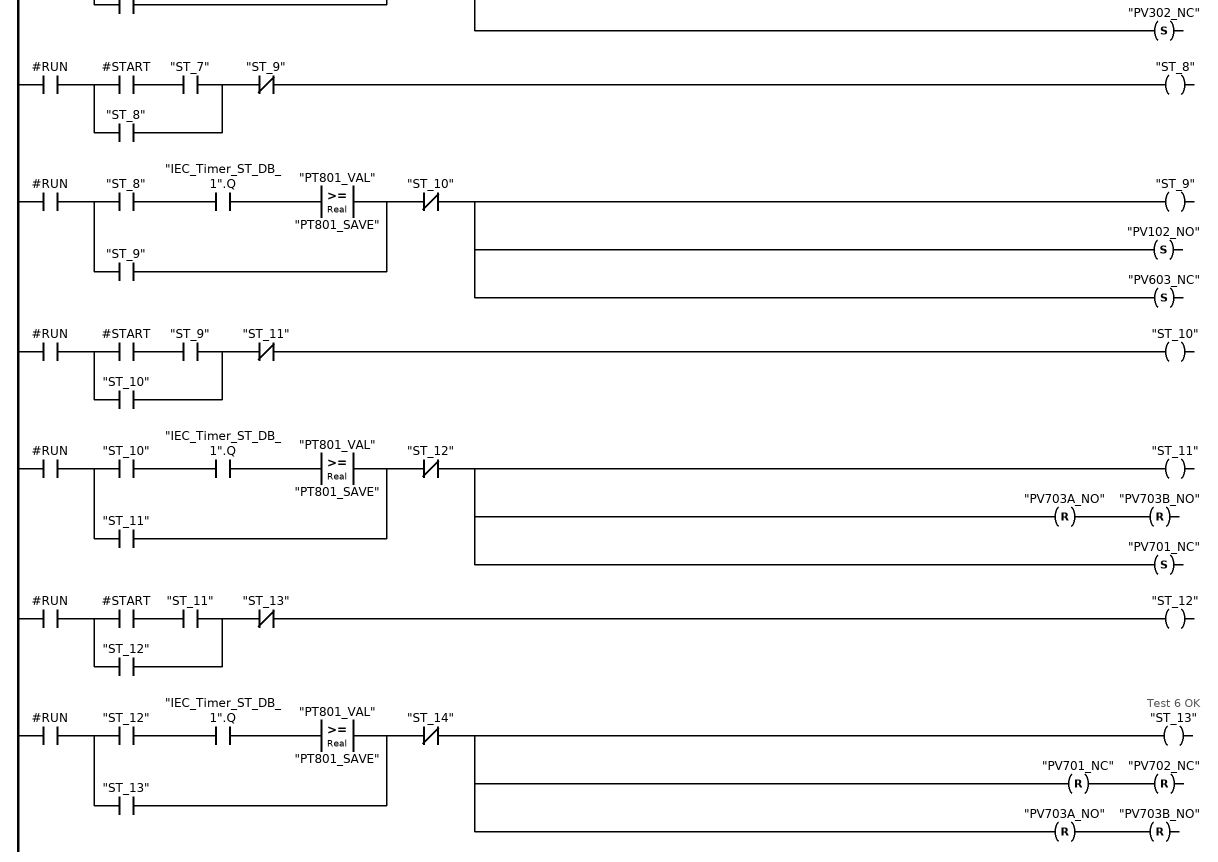
   RUNG wire#powerrail
      Contact( #RUN )
      wire#w1
      P_Contact(operand := #RUN, bit := "ST_M")
      wire#w2
      I_Contact( "ST_1" )
      I_Contact( "ST_2" )
      wire#w3
      Coil( "ST_0" )
   END_RUNG
   RUNG wire#w1
      Contact( "ST_0" )
   END_RUNG wire#w2
   RUNG wire#w3
      "ALL_VALVES_STANDBY"()
   END_RUNG
   RUNG wire#powerrail
      Contact( #RUN )
      wire#w4
      Contact( #START )
      Contact( "ST_0" )
      { S7_Templates := "SrcType := Real" } LE_Contact(in1 := "PT201_VAL", in2 := 0.0)
      { S7_Templates := "SrcType := Real" } LE_Contact(in1 := "PT401_VAL", in2 := 0.0)
      wire#w5
      I_Contact( "ST_2" )
      I_Contact( "ST_3" )
      Coil( "ST_1" )
   END_RUNG
   RUNG wire#w4
      Contact( "ST_1" )
   END_RUNG wire#w5
   RUNG wire#powerrail
      Contact( #RUN )
      wire#w6
      Contact( #START )
      Contact( "ST_1" )
      wire#w7
      I_Contact( "ST_2" )
      wire#w8
      Coil( "ST_1A" )
   END_RUNG
   RUNG wire#w6
      Contact( "ST_1A" )
   END_RUNG wire#w7
   RUNG wire#w8
      S_Coil( "PV403_NO" )
      S_Coil( "PV402_NC" )
      S_Coil( "PV602_NC" )
      S_Coil( "PV702_NC" )
   END_RUNG
   RUNG wire#w8
      Move(in := "MFC_601_MB_ADDR", out1 => "MB_DATA_MFC".MB_WRT_PARAM.MB_ADDR)
      Move(in := "MB_AD_CONTROL_MODE", out1 => "MB_DATA_MFC".MB_WRT_PARAM.DATA_ADDR)
      Move(in := "MB_VAL_CONTROL_MODE_SP_100", out1 => "MB_DATA_MFC".MB_WRT_PARAM.DATA_VAL)
   END_RUNG
   RUNG wire#powerrail
      Contact( #RUN )
      wire#w9
      Contact( "ST_1A" )
      I_Contact( "PV702_NOT_OPEN_LS" )
      wire#w10
      I_Contact( "ST_3" )
      Coil( "ST_2" )
   END_RUNG
   RUNG wire#w9
      Contact( "ST_2" )
   END_RUNG wire#w10
   RUNG wire#powerrail
      Contact( #RUN )
      wire#w11
      Contact( "ST_2" )
      Contact( "IEC_Timer_ST_DB_1".Q )
      { S7_Templates := "SrcType := Real" } GE_Contact(in1 := "PT801_VAL", in2 := "PT801_SAVE")
      wire#w12
      I_Contact( "ST_4" )
      wire#w13
      Coil( "ST_3" )
   END_RUNG
   RUNG wire#w11
      Contact( "ST_3" )
   END_RUNG wire#w12
   RUNG wire#w13
      S_Coil( "PV503_NO" )
   END_RUNG
   RUNG wire#w13
      S_Coil( "PV502_NC" )
   END_RUNG
   RUNG wire#powerrail
      Contact( #RUN )
      wire#w14
      Contact( #START )
      Contact( "ST_3" )
      wire#w15
      I_Contact( "ST_5" )
      Coil( "ST_4" )
   END_RUNG
   RUNG wire#w14
      Contact( "ST_4" )
   END_RUNG wire#w15
   RUNG wire#powerrail
      Contact( #RUN )
      wire#w16
      Contact( "ST_4" )
      Contact( "IEC_Timer_ST_DB_1".Q )
      { S7_Templates := "SrcType := Real" } GE_Contact(in1 := "PT801_VAL", in2 := "PT801_SAVE")
      wire#w17
      I_Contact( "ST_6" )
      wire#w18
      Coil( "ST_5" )
   END_RUNG
   RUNG wire#w16
      Contact( "ST_5" )
   END_RUNG wire#w17
   RUNG wire#w18
      S_Coil( "PV203_NO" )
   END_RUNG
   RUNG wire#w18
      S_Coil( "PV202_NC" )
      S_Coil( "PV601_NC" )
   END_RUNG
   RUNG wire#powerrail
      Contact( #RUN )
      wire#w19
      Contact( #START )
      Contact( "ST_5" )
      wire#w20
      I_Contact( "ST_7" )
      Coil( "ST_6" )
   END_RUNG
   RUNG wire#w19
      Contact( "ST_6" )
   END_RUNG wire#w20
   RUNG wire#powerrail
      Contact( #RUN )
      wire#w21
      Contact( "ST_6" )
      Contact( "IEC_Timer_ST_DB_1".Q )
      { S7_Templates := "SrcType := Real" } GE_Contact(in1 := "PT801_VAL", in2 := "PT801_SAVE")
      wire#w22
      I_Contact( "ST_8" )
      wire#w23
      Coil( "ST_7" )
   END_RUNG
   RUNG wire#w21
      Contact( "ST_7" )
   END_RUNG wire#w22
   RUNG wire#w23
      S_Coil( "PV303_NO" )
   END_RUNG
   RUNG wire#w23
      S_Coil( "PV302_NC" )
   END_RUNG
   RUNG wire#powerrail
      Contact( #RUN )
      wire#w24
      Contact( #START )
      Contact( "ST_7" )
      wire#w25
      I_Contact( "ST_9" )
      Coil( "ST_8" )
   END_RUNG
   RUNG wire#w24
      Contact( "ST_8" )
   END_RUNG wire#w25
   RUNG wire#powerrail
      Contact( #RUN )
      wire#w26
      Contact( "ST_8" )
      Contact( "IEC_Timer_ST_DB_1".Q )
      { S7_Templates := "SrcType := Real" } GE_Contact(in1 := "PT801_VAL", in2 := "PT801_SAVE")
      wire#w27
      I_Contact( "ST_10" )
      wire#w28
      Coil( "ST_9" )
   END_RUNG
   RUNG wire#w26
      Contact( "ST_9" )
   END_RUNG wire#w27
   RUNG wire#w28
      S_Coil( "PV102_NO" )
   END_RUNG
   RUNG wire#w28
      S_Coil( "PV603_NC" )
   END_RUNG
   RUNG wire#powerrail
      Contact( #RUN )
      wire#w29
      Contact( #START )
      Contact( "ST_9" )
      wire#w30
      I_Contact( "ST_11" )
      Coil( "ST_10" )
   END_RUNG
   RUNG wire#w29
      Contact( "ST_10" )
   END_RUNG wire#w30
   RUNG wire#powerrail
      Contact( #RUN )
      wire#w31
      Contact( "ST_10" )
      Contact( "IEC_Timer_ST_DB_1".Q )
      { S7_Templates := "SrcType := Real" } GE_Contact(in1 := "PT801_VAL", in2 := "PT801_SAVE")
      wire#w32
      I_Contact( "ST_12" )
      wire#w33
      Coil( "ST_11" )
   END_RUNG
   RUNG wire#w31
      Contact( "ST_11" )
   END_RUNG wire#w32
   RUNG wire#w33
      R_Coil( "PV703A_NO" )
      R_Coil( "PV703B_NO" )
   END_RUNG
   RUNG wire#w33
      S_Coil( "PV701_NC" )
   END_RUNG
   RUNG wire#powerrail
      Contact( #RUN )
      wire#w34
      Contact( #START )
      Contact( "ST_11" )
      wire#w35
      I_Contact( "ST_13" )
      Coil( "ST_12" )
   END_RUNG
   RUNG wire#w34
      Contact( "ST_12" )
   END_RUNG wire#w35
   RUNG wire#powerrail
      Contact( #RUN )
      wire#w36
      Contact( "ST_12" )
      Contact( "IEC_Timer_ST_DB_1".Q )
      { S7_Templates := "SrcType := Real" } GE_Contact(in1 := "PT801_VAL", in2 := "PT801_SAVE")
      wire#w37
      I_Contact( "ST_14" )
      wire#w38
      Coil( "ST_13" )   // Test 6 OK
   END_RUNG
   RUNG wire#w36
      Contact( "ST_13" )
   END_RUNG wire#w37
   RUNG wire#w38
      R_Coil( "PV701_NC" )
      R_Coil( "PV702_NC" )
   END_RUNG
   RUNG wire#w38
      R_Coil( "PV703A_NO" )
      R_Coil( "PV703B_NO" )
   END_RUNG
   // the same network as SCL:
   #_w1 := #RUN AND #RUN AND NOT "ST_M";   // rising edge of #RUN
   "ST_M" := #RUN;
   "ST_0" := (#_w1 OR (#RUN AND "ST_0")) AND NOT "ST_1" AND NOT "ST_2";
   IF "ST_0" THEN "ALL_VALVES_STANDBY"(); END_IF;
   "ST_1" := #RUN AND ((#START AND "ST_0" AND ("PT201_VAL" <= 0.0) AND ("PT401_VAL" <= 0.0)) OR "ST_1") AND NOT "ST_2" AND NOT "ST_3";
   "ST_1A" := #RUN AND ((#START AND "ST_1") OR "ST_1A") AND NOT "ST_2";
   IF "ST_1A" THEN
       "PV403_NO" := TRUE;
       "PV402_NC" := TRUE;
       "PV602_NC" := TRUE;
       "PV702_NC" := TRUE;
       "MB_DATA_MFC".MB_WRT_PARAM.MB_ADDR := "MFC_601_MB_ADDR";
       "MB_DATA_MFC".MB_WRT_PARAM.DATA_ADDR := "MB_AD_CONTROL_MODE";
       "MB_DATA_MFC".MB_WRT_PARAM.DATA_VAL := "MB_VAL_CONTROL_MODE_SP_100";
   END_IF;
   "ST_2" := #RUN AND (("ST_1A" AND NOT "PV702_NOT_OPEN_LS") OR "ST_2") AND NOT "ST_3";
   "ST_3" := #RUN AND (("ST_2" AND "IEC_Timer_ST_DB_1".Q AND ("PT801_VAL" >= "PT801_SAVE")) OR "ST_3") AND NOT "ST_4";
   IF "ST_3" THEN
       "PV503_NO" := TRUE;
       "PV502_NC" := TRUE;
   END_IF;
   "ST_4" := #RUN AND ((#START AND "ST_3") OR "ST_4") AND NOT "ST_5";
   "ST_5" := #RUN AND (("ST_4" AND "IEC_Timer_ST_DB_1".Q AND ("PT801_VAL" >= "PT801_SAVE")) OR "ST_5") AND NOT "ST_6";
   IF "ST_5" THEN
       "PV203_NO" := TRUE;
       "PV202_NC" := TRUE;
       "PV601_NC" := TRUE;
   END_IF;
   "ST_6" := #RUN AND ((#START AND "ST_5") OR "ST_6") AND NOT "ST_7";
   "ST_7" := #RUN AND (("ST_6" AND "IEC_Timer_ST_DB_1".Q AND ("PT801_VAL" >= "PT801_SAVE")) OR "ST_7") AND NOT "ST_8";
   IF "ST_7" THEN
       "PV303_NO" := TRUE;
       "PV302_NC" := TRUE;
   END_IF;
   "ST_8" := #RUN AND ((#START AND "ST_7") OR "ST_8") AND NOT "ST_9";
   "ST_9" := #RUN AND (("ST_8" AND "IEC_Timer_ST_DB_1".Q AND ("PT801_VAL" >= "PT801_SAVE")) OR "ST_9") AND NOT "ST_10";
   IF "ST_9" THEN
       "PV102_NO" := TRUE;
       "PV603_NC" := TRUE;
   END_IF;
   "ST_10" := #RUN AND ((#START AND "ST_9") OR "ST_10") AND NOT "ST_11";
   "ST_11" := #RUN AND (("ST_10" AND "IEC_Timer_ST_DB_1".Q AND ("PT801_VAL" >= "PT801_SAVE")) OR "ST_11") AND NOT "ST_12";
   IF "ST_11" THEN
       "PV703A_NO" := FALSE;
       "PV703B_NO" := FALSE;
       "PV701_NC" := TRUE;
   END_IF;
   "ST_12" := #RUN AND ((#START AND "ST_11") OR "ST_12") AND NOT "ST_13";
   "ST_13" := #RUN AND (("ST_12" AND "IEC_Timer_ST_DB_1".Q AND ("PT801_VAL" >= "PT801_SAVE")) OR "ST_13") AND NOT "ST_14";   // Test 6 OK
   IF "ST_13" THEN
       "PV701_NC" := FALSE;
       "PV702_NC" := FALSE;
       "PV703A_NO" := FALSE;
       "PV703B_NO" := FALSE;
   END_IF;
END_REGION

REGION Network 3: Process Tests
   // Tests Process Circuits  (Test #7-#9)
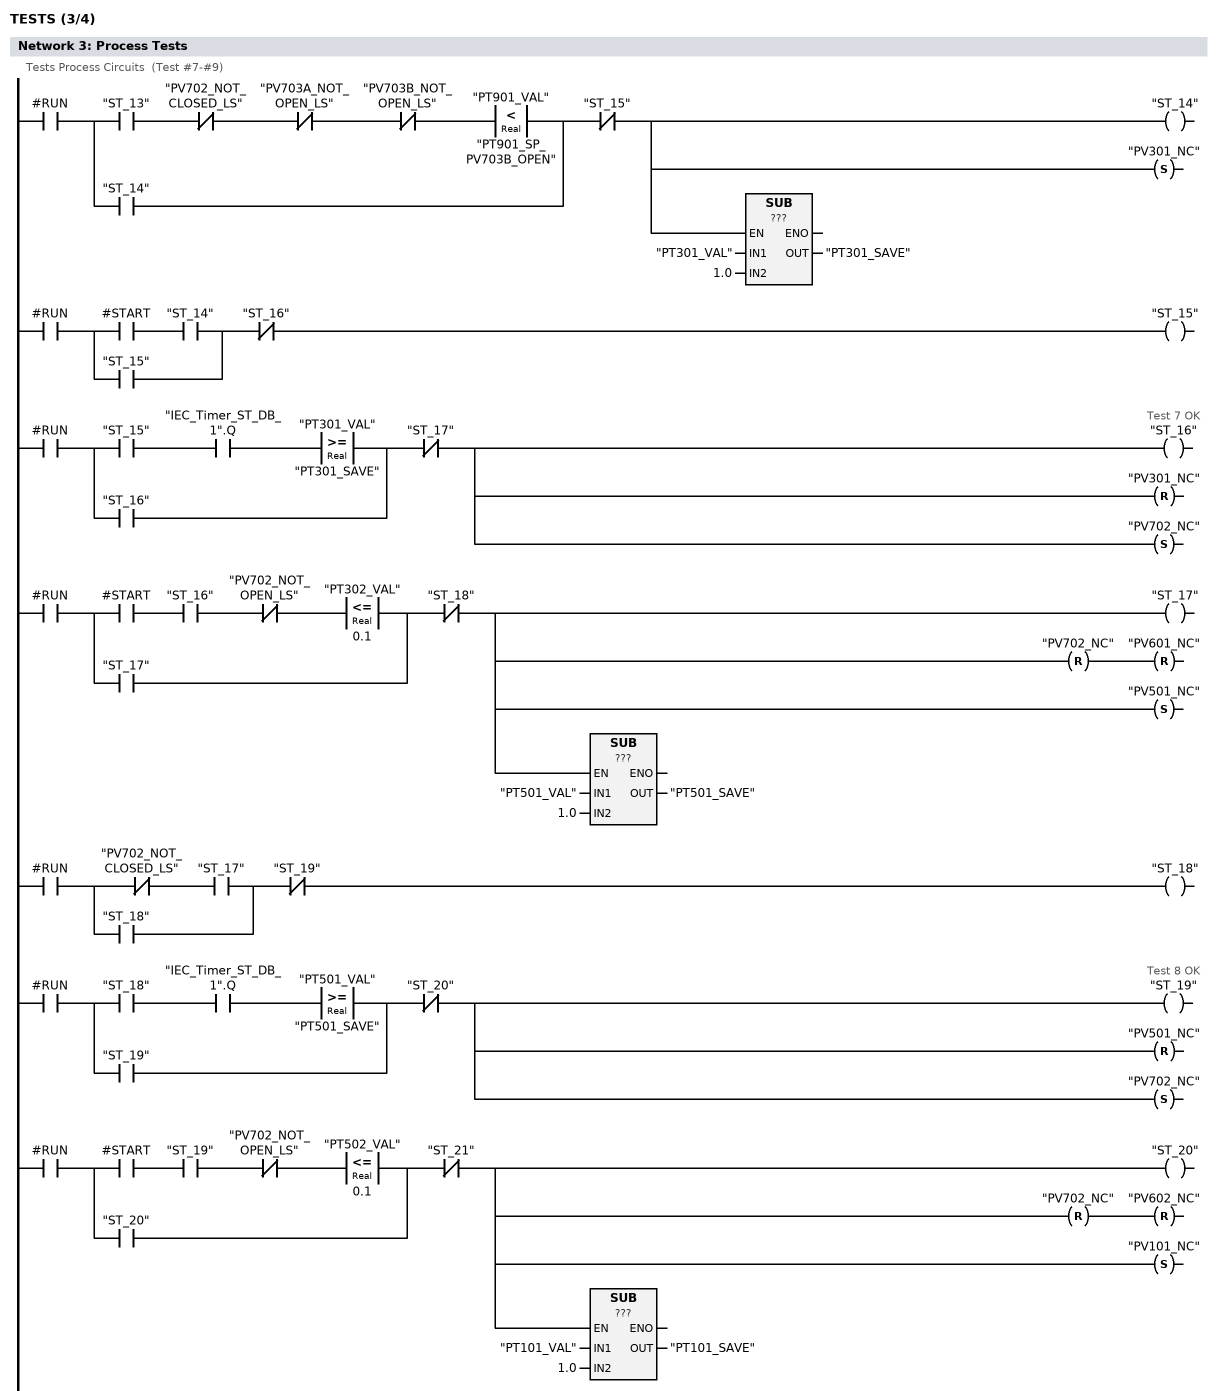
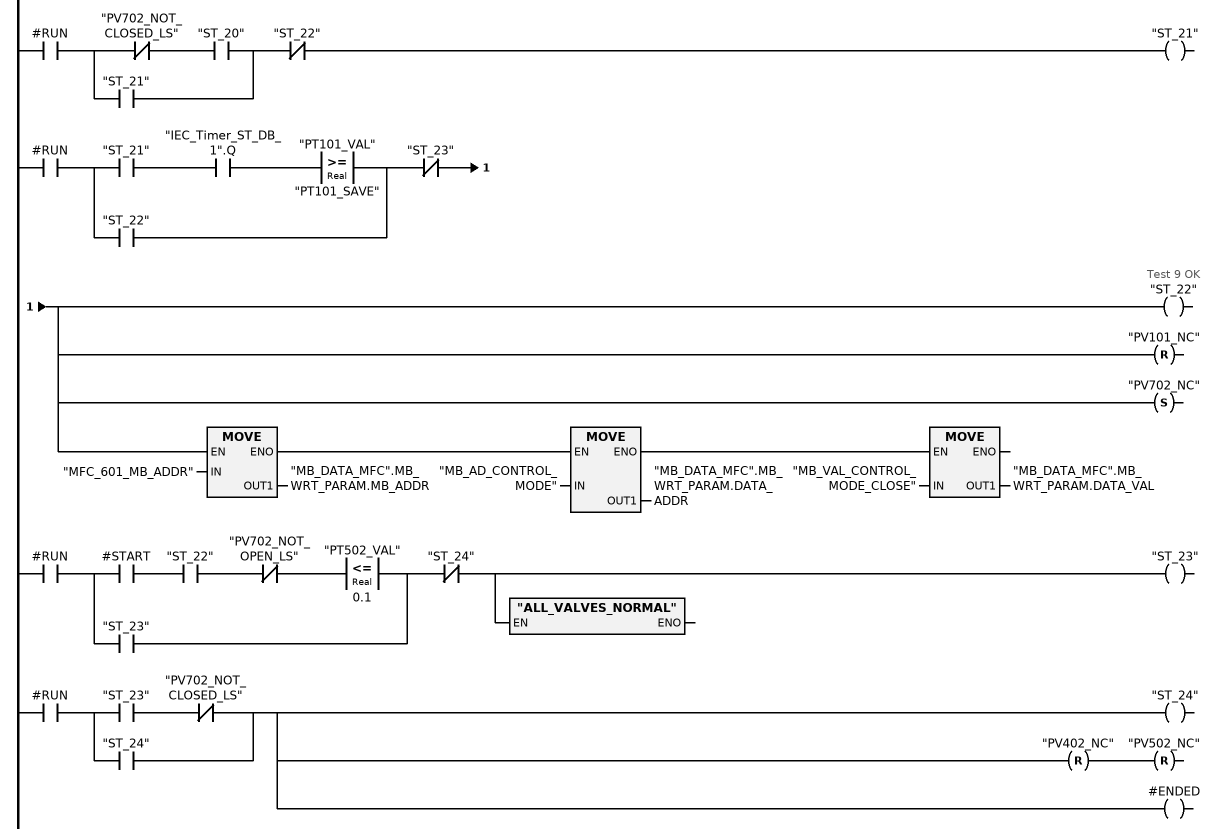
   RUNG wire#powerrail
      Contact( #RUN )
      wire#w1
      Contact( "ST_13" )
      I_Contact( "PV702_NOT_CLOSED_LS" )
      I_Contact( "PV703A_NOT_OPEN_LS" )
      I_Contact( "PV703B_NOT_OPEN_LS" )
      { S7_Templates := "SrcType := Real" } LT_Contact(in1 := "PT901_VAL", in2 := "PT901_SP_PV703B_OPEN")
      wire#w2
      I_Contact( "ST_15" )
      wire#w3
      Coil( "ST_14" )
   END_RUNG
   RUNG wire#w1
      Contact( "ST_14" )
   END_RUNG wire#w2
   RUNG wire#w3
      S_Coil( "PV301_NC" )
   END_RUNG
   RUNG wire#w3
      { S7_Templates := "SrcType := ???" } Sub(in1 := "PT301_VAL", in2 := 1.0, out => "PT301_SAVE")
   END_RUNG
   RUNG wire#powerrail
      Contact( #RUN )
      wire#w4
      Contact( #START )
      Contact( "ST_14" )
      wire#w5
      I_Contact( "ST_16" )
      Coil( "ST_15" )
   END_RUNG
   RUNG wire#w4
      Contact( "ST_15" )
   END_RUNG wire#w5
   RUNG wire#powerrail
      Contact( #RUN )
      wire#w6
      Contact( "ST_15" )
      Contact( "IEC_Timer_ST_DB_1".Q )
      { S7_Templates := "SrcType := Real" } GE_Contact(in1 := "PT301_VAL", in2 := "PT301_SAVE")
      wire#w7
      I_Contact( "ST_17" )
      wire#w8
      Coil( "ST_16" )   // Test 7 OK
   END_RUNG
   RUNG wire#w6
      Contact( "ST_16" )
   END_RUNG wire#w7
   RUNG wire#w8
      R_Coil( "PV301_NC" )
   END_RUNG
   RUNG wire#w8
      S_Coil( "PV702_NC" )
   END_RUNG
   RUNG wire#powerrail
      Contact( #RUN )
      wire#w9
      Contact( #START )
      Contact( "ST_16" )
      I_Contact( "PV702_NOT_OPEN_LS" )
      { S7_Templates := "SrcType := Real" } LE_Contact(in1 := "PT302_VAL", in2 := 0.1)
      wire#w10
      I_Contact( "ST_18" )
      wire#w11
      Coil( "ST_17" )
   END_RUNG
   RUNG wire#w9
      Contact( "ST_17" )
   END_RUNG wire#w10
   RUNG wire#w11
      R_Coil( "PV702_NC" )
      R_Coil( "PV601_NC" )
   END_RUNG
   RUNG wire#w11
      S_Coil( "PV501_NC" )
   END_RUNG
   RUNG wire#w11
      { S7_Templates := "SrcType := ???" } Sub(in1 := "PT501_VAL", in2 := 1.0, out => "PT501_SAVE")
   END_RUNG
   RUNG wire#powerrail
      Contact( #RUN )
      wire#w12
      I_Contact( "PV702_NOT_CLOSED_LS" )
      Contact( "ST_17" )
      wire#w13
      I_Contact( "ST_19" )
      Coil( "ST_18" )
   END_RUNG
   RUNG wire#w12
      Contact( "ST_18" )
   END_RUNG wire#w13
   RUNG wire#powerrail
      Contact( #RUN )
      wire#w14
      Contact( "ST_18" )
      Contact( "IEC_Timer_ST_DB_1".Q )
      { S7_Templates := "SrcType := Real" } GE_Contact(in1 := "PT501_VAL", in2 := "PT501_SAVE")
      wire#w15
      I_Contact( "ST_20" )
      wire#w16
      Coil( "ST_19" )   // Test 8 OK
   END_RUNG
   RUNG wire#w14
      Contact( "ST_19" )
   END_RUNG wire#w15
   RUNG wire#w16
      R_Coil( "PV501_NC" )
   END_RUNG
   RUNG wire#w16
      S_Coil( "PV702_NC" )
   END_RUNG
   RUNG wire#powerrail
      Contact( #RUN )
      wire#w17
      Contact( #START )
      Contact( "ST_19" )
      I_Contact( "PV702_NOT_OPEN_LS" )
      { S7_Templates := "SrcType := Real" } LE_Contact(in1 := "PT502_VAL", in2 := 0.1)
      wire#w18
      I_Contact( "ST_21" )
      wire#w19
      Coil( "ST_20" )
   END_RUNG
   RUNG wire#w17
      Contact( "ST_20" )
   END_RUNG wire#w18
   RUNG wire#w19
      R_Coil( "PV702_NC" )
      R_Coil( "PV602_NC" )
   END_RUNG
   RUNG wire#w19
      S_Coil( "PV101_NC" )
   END_RUNG
   RUNG wire#w19
      { S7_Templates := "SrcType := ???" } Sub(in1 := "PT101_VAL", in2 := 1.0, out => "PT101_SAVE")
   END_RUNG
   RUNG wire#powerrail
      Contact( #RUN )
      wire#w20
      I_Contact( "PV702_NOT_CLOSED_LS" )
      Contact( "ST_20" )
      wire#w21
      I_Contact( "ST_22" )
      Coil( "ST_21" )
   END_RUNG
   RUNG wire#w20
      Contact( "ST_21" )
   END_RUNG wire#w21
   RUNG wire#powerrail
      Contact( #RUN )
      wire#w22
      Contact( "ST_21" )
      Contact( "IEC_Timer_ST_DB_1".Q )
      { S7_Templates := "SrcType := Real" } GE_Contact(in1 := "PT101_VAL", in2 := "PT101_SAVE")
      wire#w23
      I_Contact( "ST_23" )
      wire#w24
      Coil( "ST_22" )   // Test 9 OK
   END_RUNG
   RUNG wire#w22
      Contact( "ST_22" )
   END_RUNG wire#w23
   RUNG wire#w24
      R_Coil( "PV101_NC" )
   END_RUNG
   RUNG wire#w24
      S_Coil( "PV702_NC" )
   END_RUNG
   RUNG wire#w24
      Move(in := "MFC_601_MB_ADDR", out1 => "MB_DATA_MFC".MB_WRT_PARAM.MB_ADDR)
      Move(in := "MB_AD_CONTROL_MODE", out1 => "MB_DATA_MFC".MB_WRT_PARAM.DATA_ADDR)
      Move(in := "MB_VAL_CONTROL_MODE_CLOSE", out1 => "MB_DATA_MFC".MB_WRT_PARAM.DATA_VAL)
   END_RUNG
   RUNG wire#powerrail
      Contact( #RUN )
      wire#w25
      Contact( #START )
      Contact( "ST_22" )
      I_Contact( "PV702_NOT_OPEN_LS" )
      { S7_Templates := "SrcType := Real" } LE_Contact(in1 := "PT502_VAL", in2 := 0.1)
      wire#w26
      I_Contact( "ST_24" )
      wire#w27
      Coil( "ST_23" )
   END_RUNG
   RUNG wire#w25
      Contact( "ST_23" )
   END_RUNG wire#w26
   RUNG wire#w27
      "ALL_VALVES_NORMAL"()
   END_RUNG
   RUNG wire#powerrail
      Contact( #RUN )
      wire#w28
      Contact( "ST_23" )
      I_Contact( "PV702_NOT_CLOSED_LS" )
      wire#w29
      Coil( "ST_24" )
   END_RUNG
   RUNG wire#w28
      Contact( "ST_24" )
   END_RUNG wire#w29
   RUNG wire#w29
      R_Coil( "PV402_NC" )
      R_Coil( "PV502_NC" )
   END_RUNG
   RUNG wire#w29
      Coil( #ENDED )
   END_RUNG
   // the same network as SCL:
   "ST_14" := #RUN AND (("ST_13" AND NOT "PV702_NOT_CLOSED_LS" AND NOT "PV703A_NOT_OPEN_LS" AND NOT "PV703B_NOT_OPEN_LS" AND ("PT901_VAL" < "PT901_SP_PV703B_OPEN")) OR "ST_14") AND NOT "ST_15";
   IF "ST_14" THEN
       "PV301_NC" := TRUE;
       "PT301_SAVE" := "PT301_VAL" - 1.0;
   END_IF;
   "ST_15" := #RUN AND ((#START AND "ST_14") OR "ST_15") AND NOT "ST_16";
   "ST_16" := #RUN AND (("ST_15" AND "IEC_Timer_ST_DB_1".Q AND ("PT301_VAL" >= "PT301_SAVE")) OR "ST_16") AND NOT "ST_17";   // Test 7 OK
   IF "ST_16" THEN
       "PV301_NC" := FALSE;
       "PV702_NC" := TRUE;
   END_IF;
   "ST_17" := #RUN AND ((#START AND "ST_16" AND NOT "PV702_NOT_OPEN_LS" AND ("PT302_VAL" <= 0.1)) OR "ST_17") AND NOT "ST_18";
   IF "ST_17" THEN
       "PV702_NC" := FALSE;
       "PV601_NC" := FALSE;
       "PV501_NC" := TRUE;
       "PT501_SAVE" := "PT501_VAL" - 1.0;
   END_IF;
   "ST_18" := #RUN AND ((NOT "PV702_NOT_CLOSED_LS" AND "ST_17") OR "ST_18") AND NOT "ST_19";
   "ST_19" := #RUN AND (("ST_18" AND "IEC_Timer_ST_DB_1".Q AND ("PT501_VAL" >= "PT501_SAVE")) OR "ST_19") AND NOT "ST_20";   // Test 8 OK
   IF "ST_19" THEN
       "PV501_NC" := FALSE;
       "PV702_NC" := TRUE;
   END_IF;
   "ST_20" := #RUN AND ((#START AND "ST_19" AND NOT "PV702_NOT_OPEN_LS" AND ("PT502_VAL" <= 0.1)) OR "ST_20") AND NOT "ST_21";
   IF "ST_20" THEN
       "PV702_NC" := FALSE;
       "PV602_NC" := FALSE;
       "PV101_NC" := TRUE;
       "PT101_SAVE" := "PT101_VAL" - 1.0;
   END_IF;
   "ST_21" := #RUN AND ((NOT "PV702_NOT_CLOSED_LS" AND "ST_20") OR "ST_21") AND NOT "ST_22";
   "ST_22" := #RUN AND (("ST_21" AND "IEC_Timer_ST_DB_1".Q AND ("PT101_VAL" >= "PT101_SAVE")) OR "ST_22") AND NOT "ST_23";   // Test 9 OK
   IF "ST_22" THEN
       "PV101_NC" := FALSE;
       "PV702_NC" := TRUE;
       "MB_DATA_MFC".MB_WRT_PARAM.MB_ADDR := "MFC_601_MB_ADDR";
       "MB_DATA_MFC".MB_WRT_PARAM.DATA_ADDR := "MB_AD_CONTROL_MODE";
       "MB_DATA_MFC".MB_WRT_PARAM.DATA_VAL := "MB_VAL_CONTROL_MODE_CLOSE";
   END_IF;
   "ST_23" := #RUN AND ((#START AND "ST_22" AND NOT "PV702_NOT_OPEN_LS" AND ("PT502_VAL" <= 0.1)) OR "ST_23") AND NOT "ST_24";
   IF "ST_23" THEN "ALL_VALVES_NORMAL"(); END_IF;
   "ST_24" := #RUN AND (("ST_23" AND NOT "PV702_NOT_CLOSED_LS") OR "ST_24");
   IF "ST_24" THEN
       "PV402_NC" := FALSE;
       "PV502_NC" := FALSE;
   END_IF;
   #ENDED := "ST_24";
END_REGION

REGION Network 4
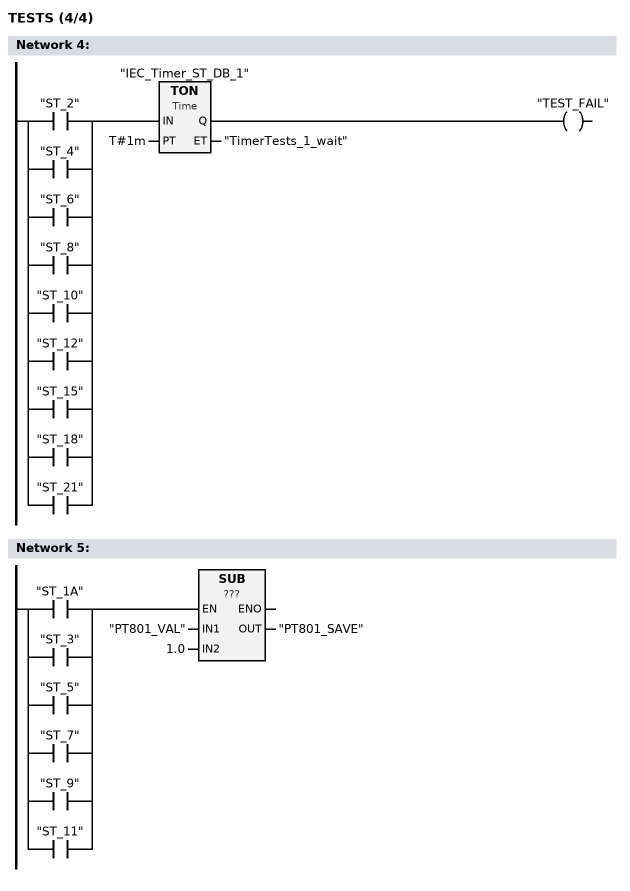
   "IEC_Timer_ST_DB_1".TON(IN := "ST_2" OR "ST_4" OR "ST_6" OR "ST_8" OR "ST_10" OR "ST_12" OR "ST_15" OR "ST_18" OR "ST_21",
                           PT := T#1m,
                           ET => "TimerTests_1_wait");
   "TEST_FAIL" := "IEC_Timer_ST_DB_1".Q;
END_REGION

REGION Network 5
   RUNG wire#powerrail
      Contact( "ST_1A" )
      wire#w1
      { S7_Templates := "SrcType := ???" } Sub(in1 := "PT801_VAL", in2 := 1.0, out => "PT801_SAVE")
   END_RUNG
   RUNG wire#powerrail
      Contact( "ST_3" )
   END_RUNG wire#w1
   RUNG wire#powerrail
      Contact( "ST_5" )
   END_RUNG wire#w1
   RUNG wire#powerrail
      Contact( "ST_7" )
   END_RUNG wire#w1
   RUNG wire#powerrail
      Contact( "ST_9" )
   END_RUNG wire#w1
   RUNG wire#powerrail
      Contact( "ST_11" )
   END_RUNG wire#w1
   // the same network as SCL:
   IF "ST_1A" OR "ST_3" OR "ST_5" OR "ST_7" OR "ST_9" OR "ST_11" THEN
       "PT801_SAVE" := "PT801_VAL" - 1.0;
   END_IF;
END_REGION
END_FUNCTION

FUNCTION "ETAPA_9" : Void   // FC11, LAD
TITLE = ETAPA 9 - EXAUSTÃO
{ S7_Optimized_Access := 'FALSE' }
VERSION : 0.1
BEGIN

REGION Network 1
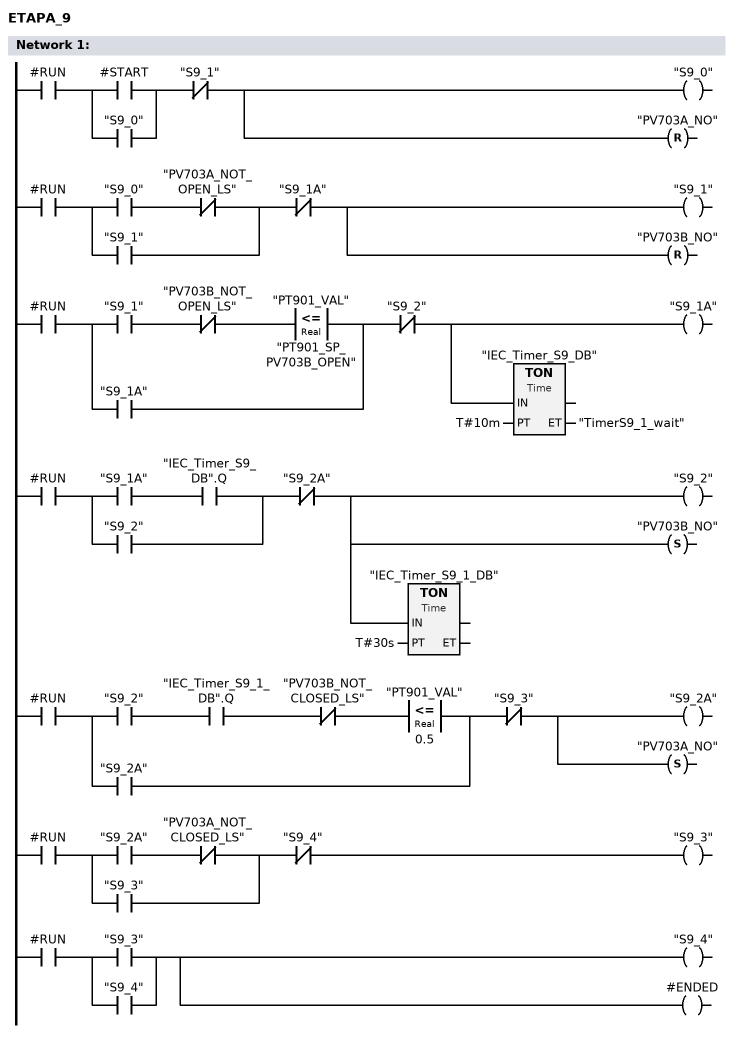
   "S9_0" := #RUN AND (#START OR "S9_0") AND NOT "S9_1";
   IF "S9_0" THEN "PV703A_NO" := FALSE; END_IF;
   "S9_1" := #RUN AND (("S9_0" AND NOT "PV703A_NOT_OPEN_LS") OR "S9_1") AND NOT "S9_1A";
   IF "S9_1" THEN "PV703B_NO" := FALSE; END_IF;
   "S9_1A" := #RUN AND (("S9_1" AND NOT "PV703B_NOT_OPEN_LS" AND ("PT901_VAL" <= "PT901_SP_PV703B_OPEN")) OR "S9_1A") AND NOT "S9_2";
   "IEC_Timer_S9_DB".TON(IN := "S9_1A", PT := T#10m, ET => "TimerS9_1_wait");
   "S9_2" := #RUN AND (("S9_1A" AND "IEC_Timer_S9_DB".Q) OR "S9_2") AND NOT "S9_2A";
   IF "S9_2" THEN "PV703B_NO" := TRUE; END_IF;
   "IEC_Timer_S9_1_DB".TON(IN := "S9_2", PT := T#30s);
   "S9_2A" := #RUN AND (("S9_2" AND "IEC_Timer_S9_1_DB".Q AND NOT "PV703B_NOT_CLOSED_LS" AND ("PT901_VAL" <= 0.5)) OR "S9_2A") AND NOT "S9_3";
   IF "S9_2A" THEN "PV703A_NO" := TRUE; END_IF;
   "S9_3" := #RUN AND (("S9_2A" AND NOT "PV703A_NOT_CLOSED_LS") OR "S9_3") AND NOT "S9_4";
   "S9_4" := #RUN AND ("S9_3" OR "S9_4");
   #ENDED := "S9_4";
END_REGION
END_FUNCTION

FUNCTION "MB_Cyclic_Read" : Void   // FC12, LAD
{ S7_Optimized_Access := 'FALSE' }
VERSION : 0.1
   VAR_TEMP   // added for the SCL form of the ladder/FBD networks
      _w1 : Bool;
   END_VAR
BEGIN

REGION Network 1
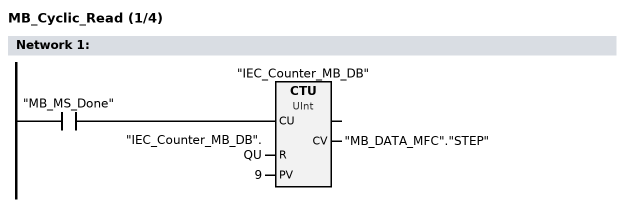
   "IEC_Counter_MB_DB".CTU(CU := "MB_MS_Done", R := "IEC_Counter_MB_DB".QU, PV := 9, CV => "MB_DATA_MFC"."STEP");
END_REGION

REGION Network 2
   // MODBUS MASTER Cyclic Read
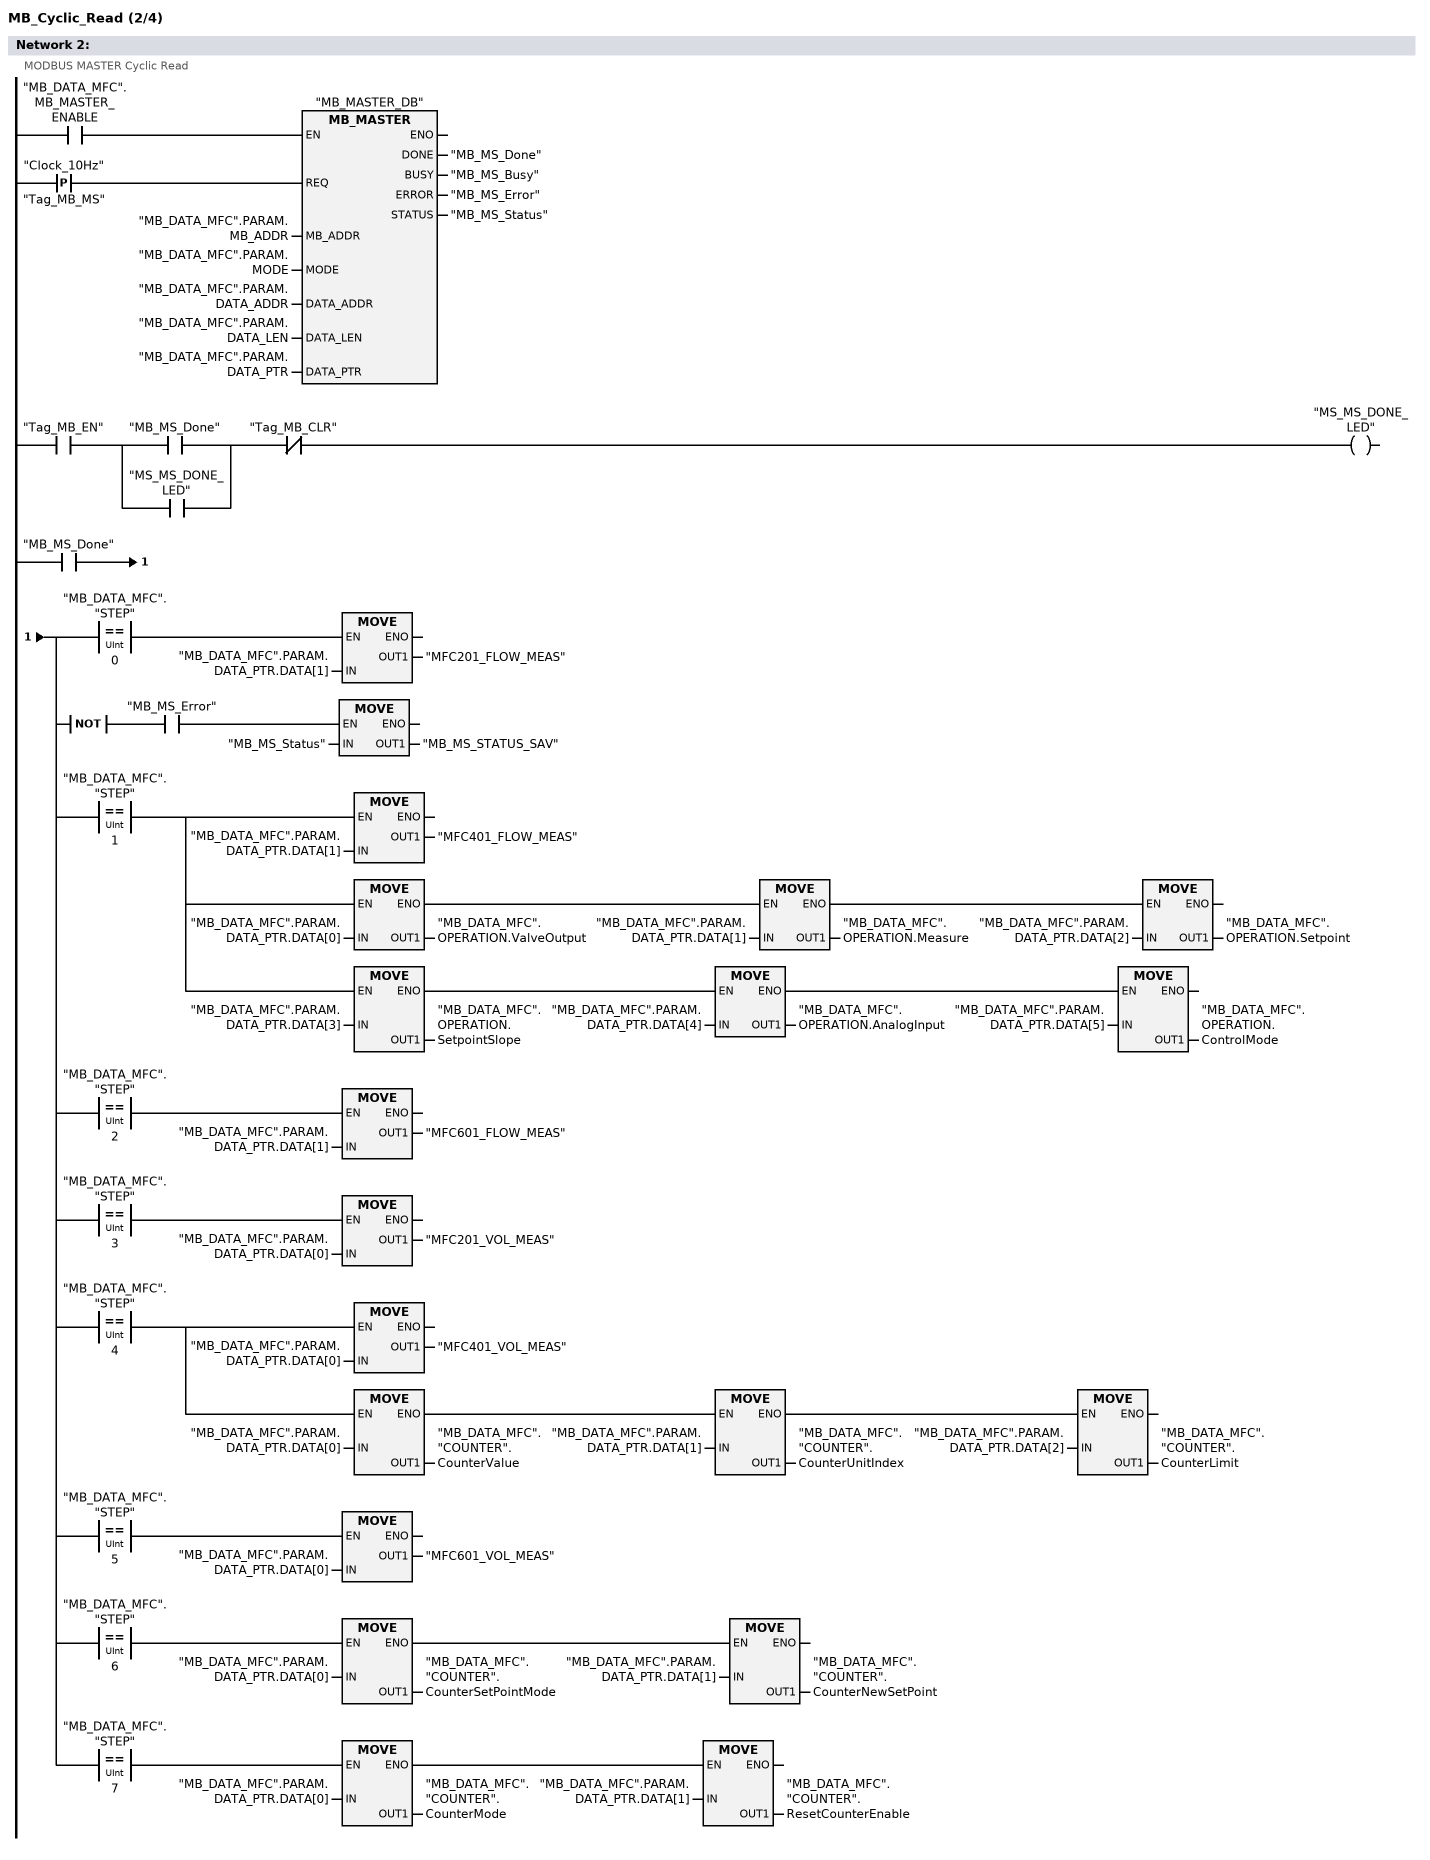
   #_w1 := "Clock_10Hz" AND NOT "Tag_MB_MS";   // rising edge of "Clock_10Hz"
   "Tag_MB_MS" := "Clock_10Hz";
   IF "MB_DATA_MFC".MB_MASTER_ENABLE THEN
       "MB_MASTER_DB"(REQ := #_w1,   // MB_MASTER
                      MB_ADDR := "MB_DATA_MFC".PARAM.MB_ADDR,
                      MODE := "MB_DATA_MFC".PARAM.MODE,
                      DATA_ADDR := "MB_DATA_MFC".PARAM.DATA_ADDR,
                      DATA_LEN := "MB_DATA_MFC".PARAM.DATA_LEN,
                      DATA_PTR := "MB_DATA_MFC".PARAM.DATA_PTR,
                      DONE => "MB_MS_Done",
                      BUSY => "MB_MS_Busy",
                      ERROR => "MB_MS_Error",
                      STATUS => "MB_MS_Status");
   END_IF;
   "MS_MS_DONE_LED" := "Tag_MB_EN" AND ("MB_MS_Done" OR "MS_MS_DONE_LED") AND NOT "Tag_MB_CLR";
   IF "MB_MS_Done" AND ("MB_DATA_MFC"."STEP" = 0) THEN
       "MFC201_FLOW_MEAS" := "MB_DATA_MFC".PARAM.DATA_PTR.DATA[1];
   END_IF;
   IF NOT "MB_MS_Done" AND "MB_MS_Error" THEN "MB_MS_STATUS_SAV" := "MB_MS_Status"; END_IF;
   IF "MB_MS_Done" AND ("MB_DATA_MFC"."STEP" = 1) THEN
       "MFC401_FLOW_MEAS" := "MB_DATA_MFC".PARAM.DATA_PTR.DATA[1];
       "MB_DATA_MFC".OPERATION.ValveOutput := "MB_DATA_MFC".PARAM.DATA_PTR.DATA[0];
       "MB_DATA_MFC".OPERATION.Measure := "MB_DATA_MFC".PARAM.DATA_PTR.DATA[1];
       "MB_DATA_MFC".OPERATION.Setpoint := "MB_DATA_MFC".PARAM.DATA_PTR.DATA[2];
       "MB_DATA_MFC".OPERATION.SetpointSlope := "MB_DATA_MFC".PARAM.DATA_PTR.DATA[3];
       "MB_DATA_MFC".OPERATION.AnalogInput := "MB_DATA_MFC".PARAM.DATA_PTR.DATA[4];
       "MB_DATA_MFC".OPERATION.ControlMode := "MB_DATA_MFC".PARAM.DATA_PTR.DATA[5];
   END_IF;
   IF "MB_MS_Done" AND ("MB_DATA_MFC"."STEP" = 2) THEN
       "MFC601_FLOW_MEAS" := "MB_DATA_MFC".PARAM.DATA_PTR.DATA[1];
   END_IF;
   IF "MB_MS_Done" AND ("MB_DATA_MFC"."STEP" = 3) THEN
       "MFC201_VOL_MEAS" := "MB_DATA_MFC".PARAM.DATA_PTR.DATA[0];
   END_IF;
   IF "MB_MS_Done" AND ("MB_DATA_MFC"."STEP" = 4) THEN
       "MFC401_VOL_MEAS" := "MB_DATA_MFC".PARAM.DATA_PTR.DATA[0];
       "MB_DATA_MFC"."COUNTER".CounterValue := "MB_DATA_MFC".PARAM.DATA_PTR.DATA[0];
       "MB_DATA_MFC"."COUNTER".CounterUnitIndex := "MB_DATA_MFC".PARAM.DATA_PTR.DATA[1];
       "MB_DATA_MFC"."COUNTER".CounterLimit := "MB_DATA_MFC".PARAM.DATA_PTR.DATA[2];
   END_IF;
   IF "MB_MS_Done" AND ("MB_DATA_MFC"."STEP" = 5) THEN
       "MFC601_VOL_MEAS" := "MB_DATA_MFC".PARAM.DATA_PTR.DATA[0];
   END_IF;
   IF "MB_MS_Done" AND ("MB_DATA_MFC"."STEP" = 6) THEN
       "MB_DATA_MFC"."COUNTER".CounterSetPointMode := "MB_DATA_MFC".PARAM.DATA_PTR.DATA[0];
       "MB_DATA_MFC"."COUNTER".CounterNewSetPoint := "MB_DATA_MFC".PARAM.DATA_PTR.DATA[1];
   END_IF;
   IF "MB_MS_Done" AND ("MB_DATA_MFC"."STEP" = 7) THEN
       "MB_DATA_MFC"."COUNTER".CounterMode := "MB_DATA_MFC".PARAM.DATA_PTR.DATA[0];
       "MB_DATA_MFC"."COUNTER".ResetCounterEnable := "MB_DATA_MFC".PARAM.DATA_PTR.DATA[1];
   END_IF;
END_REGION

REGION Network 3
   // Read address on each cycle